// TIA Portal project "FK_PiPl" (V16)
// Lehrlingsprojekt

(* hardware
DEVICE "ET 200SP-Station_1"  ET 200SP-Station
   slot 0: "Baugruppenträger_0"  Rack  6ES5 710-8MAx1
   slot 1: "-20KF1"  CPU 1512SP F-1 PN  6ES7 512-1SK01-0AB0  V2.8
      slot 32768: "PROFINET-Schnittstelle_1"  X1
         slot 32771: "Port_3"  X1 P3
   slot 2: "-20KF5"  F-DI 8x24VDC HF  6ES7 136-6BA00-0CA0  V1.0
      slot 1: "-20KF5"  F-DI 8x24VDC HF
   slot 3: "-20KF6"  F-DQ 8x24VDC/0.5A PP HF  6ES7 136-6DC00-0CA0  V1.0
      slot 1: "-20KF6"  F-DQ 8x24VDC/0.5A PP HF
   slot 4: "-21KF1"  DI 16x24VDC ST  6ES7 131-6BH01-0BA0  V0.0
      slot 1: "-21KF1"  DI 16x24VDC ST
   slot 5: "-21KF4"  DQ 16x24VDC/0.5A ST  6ES7 132-6BH01-0BA0  V0.0
      slot 1: "-21KF4"  DQ 16x24VDC/0.5A ST
   slot 6: "-22KF1"  AI 2xU/I 2-,4-wire HS  6ES7 134-6HB00-0DA1  V2.0
      slot 1: "-22KF1"  AI 2xU/I 2-,4-wire HS
   slot 7: "-22KF3"  AQ 2xU ST  6ES7 135-6FB00-0BA1  V1.0
      slot 1: "-22KF3"  AQ 2xU ST
   slot 8: "Servermodul_1"  Server module  6ES7 193-6PA00-0AA0  V1.1
      slot 1: "Servermodul_1"  Server module
   slot 127: "BA 2xRJ45"  BA 2xRJ45  6ES7 193-6AR00-0AA0  V0.0
      slot 32769: "Port_1"  X1 P1  6ES7 193-6AR00-0AA0
      slot 32770: "Port_2"  X1 P2  6ES7 193-6AR00-0AA0
DEVICE "HMI_1"  KTP400 Comfort
   slot 0: "HMI_1"  KTP400 Comfort  6AV2 124-2DC01-0AX0  16.0.0.0
   slot 1: "HMI_RT_1"  KTP400 Comfort  6AV2 124-2DC01-0AX0  16.0.0.0
   slot 5: "HMI_1.IE_CP_1"  PROFINET Interface  16.0.0.0
      slot 1: "PROFINET Schnittstelle_1"  PROFINET Interface
         slot 1: "Port_1"  Port
   slot 7: "HMI_1.MPI/DP_CP_1"  MPI/DP Interface  16.0.0.0
*)

// ===== PLC "-20KF1"  CPU 1512SP F-1 PN =====
// protected blocks, not shown: "Datenbaustein_2", "Main_Safety_RTG1", "Main_Safety_RTG1_DB", "Safety_Variabeln"

VAR_GLOBAL   // PLC tag table "Standard-Variablentabelle"
   "Speicher_Start" AT %M4.0 : Bool;
   "Speicher_Vereinzelner" AT %M4.1 : Bool;
   "Speicher_Teil_Bereit" AT %M4.2 : Bool;
   "Flanke_Teil_Bereit" AT %M4.3 : Bool;
   "Deckel_Drauf" AT %M4.4 : Bool;
   "Sauger_an" AT %M4.6 : Bool;
   "Sauger_Runter" AT %M4.7 : Bool;
   "Schlitten_Ausfahren" AT %M5.0 : Bool;
   "Flanke_Schltten_Ausgefahren" AT %M5.1 : Bool;
   "Speicher_Schlitten_Ausgefahren" AT %M5.2 : Bool;
   "Flanke_Schlitten" AT %M5.3 : Bool;
   "Flanke_Teil" AT %M5.4 : Bool;
   "Speicher_Sauger_aktivierung" AT %M5.5 : Bool;
   "Teil_Fertig" AT %M5.6 : Bool;
   "Speicher_kein_Deckel" AT %M5.7 : Bool;
   "Start/Stop Auto" AT %M6.0 : Bool;
   "Flanke_Dekel" AT %M6.1 : Bool;
   "Merker_Flanke_kein_Deckel" AT %M6.2 : Bool;
   "Speicher_Rückstau" AT %M6.3 : Bool;
   "Förderband-vor_Speicher" AT %M4.5 : Bool;
   "Förderband_Zurück_Speicher" AT %M6.4 : Bool;
   "Start/Stop Hand" AT %M6.5 : Bool;
   "Druck_Sensor" AT %EW272 : Word;
   "Druck_Zwischenwert1" AT %MD100 : Real;
   "Druck_Zwischenwert2" AT %MD104 : Real;
   "Druck_Zwischenwert3" AT %MW108 : Int;
   "Druck_Zugross" AT %M6.6 : Bool;
   "Druck_Zuklein" AT %M6.7 : Bool;
   "Flanke p Man/Aut" AT %M7.0 : Bool;
   "Flanke n Man/Aut" AT %M7.1 : Bool;
   "Flanke Merker n Man/Aut" AT %M7.2 : Bool;
   "Flanke Merker p Man/Aut" AT %M7.3 : Bool;
   "Reset Man/Aut" AT %M7.4 : Bool;
END_VAR

VAR_GLOBAL   // PLC tag table "Systemflags"
   "System_Byte" AT %MB1 : Byte;   // Byte System
   "ME_PLC_First_Scan_Bit" AT %M1.0 : Bool;   // PLC First Scan Bit
   "ME_PLC_DiagStatusUpdate" AT %M1.1 : Bool;   // PLC Diagnostic Status Update
   "ME_PLC_TRUE" AT %M1.2 : Bool;   // PLC TRUE
   "ME_PLC_FALSE" AT %M1.3 : Bool;   // PLC FALSE
   "Clock_Byte" AT %MB50 : Byte;   // Byte PLC Clock
   "ME_PLC_Clock_0.1s" AT %M50.0 : Bool;   // PLC Clock 0.1s (10Hz )
   "ME_PLC_Clock_0.2s" AT %M50.1 : Bool;   // PLC Clock 0.2s (5Hz )
   "ME_PLC_Clock_0.4s" AT %M50.2 : Bool;   // PLC Clock 0.4s (2.5Hz )
   "ME_PLC_Clock_0.5s" AT %M50.3 : Bool;   // PLC Clock 0.5s (2Hz )
   "ME_PLC_Clock_0.8s" AT %M50.4 : Bool;   // PLC Clock 0.8s (1.25Hz )
   "ME_PLC_Clock_1.0s" AT %M50.5 : Bool;   // PLC Clock 1s (1Hz)
   "ME_PLC_Clock_1.6s" AT %M50.6 : Bool;   // PLC Clock 1.6s (0.625Hz )
   "ME_PLC_Clock_2.0s" AT %M50.7 : Bool;   // PLC Clock 2s (0.5Hz )
   "ME_PLC_FC_Test" AT %M2.0 : Bool;   // Testing Frequency Converters
   "ME_PLC_TRUE_to_do" AT %M2.2 : Bool;   // PLC TRUE to do
   "ME_PLC_FALSE_to_do" AT %M2.3 : Bool;   // PLC FALSE to do
   "ME_PLC_Led_Error" AT %M2.4 : Bool;   // PLC LED Error
   "ME_PLC_Led_Maint" AT %M2.5 : Bool;   // PLC LED Maintenance
   "ME_PLC_Startup_Rst" AT %M2.6 : Bool;   // PLC LED Startup Reset
   "ME_PLC_First_Scan_Bit_FC" AT %M2.1 : Bool;   // Call Frequency Converters
END_VAR

VAR_GLOBAL   // PLC tag table "IO-Pick&Placer"
   "CC_KF_FbEStop" AT %E0.0 : Bool;   // Rückmeldung Freigabe Not-Halt (81KF8)
   "PPTR_BG_InletPart" AT %E0.1 : Bool;   // Transportband Werkstück am Bandanfang (100BG1)
   "PPTR_BG_PartAtSep" AT %E0.2 : Bool;   // Transportband Werkstück am Vereinzeler (100BG2)
   "PPTR_BG_BackupPart" AT %E0.3 : Bool;   // Transportband Werkstück beim Bandende (100BG3)
   "PIPL_BG_CarrierRetracted" AT %E0.4 : Bool;   // Pick&Placer Schlitten eingefahren (120BG1)
   "PIPL_BG_CarrierExtended" AT %E0.5 : Bool;   // Pick&Placer Schlitten ausgefahren (120BG2)
   "PIPL_BG_SuctTop" AT %E0.6 : Bool;   // Pick&Placer Sauger oben (120BG3)
   "PIPL_BP_PartSuckedOn" AT %E0.7 : Bool;   // Pick&Placer Werkstück angesaugt (120PB4)
   "PIPL_Pa_SF_Reset" AT %E1.0 : Bool;   // Pick&Placer Bedienstelle Reset (160SF2)
   "PIPL_Pa_SF_Start" AT %E1.1 : Bool;   // Pick&Placer Bedienstelle Start (160SF3)
   "PIPL_Pa_SF_Stop" AT %E1.2 : Bool;   // Pick&Placer Bedienstelle Stop (160SF4)
   "PIPL_Pa_SF_ManAuto" AT %E1.3 : Bool;   // Pick&Placer Bedienstelle Manual - Auto (160SF5)
   "CC_Spare_I1.4" AT %E1.4 : Bool;   // Spare
   "CC_Spare_I1.5" AT %E1.5 : Bool;   // Spare
   "CC_Spare_I1.6" AT %E1.6 : Bool;   // Spare
   "CC_Spare_I1.7" AT %E1.7 : Bool;   // Spare
   "PPTR_MB_SeparatorExtend" AT %A0.0 : Bool;   // Transportband Vereinzeler ausfahren (105MB8)
   "PIPL_SC_Green" AT %A0.1 : Bool;   // Pick&Placer Turmleuchte grün (130PF1)
   "PIPL_SC_Yellow" AT %A0.2 : Bool;   // Pick&Placer Turmleuchte gelb (130PF1)
   "PIPL_SC_Red" AT %A0.3 : Bool;   // Pick&Placer Turmleuchte rot (130PF1)
   "PIPL_MB_CarrierExtend" AT %A0.4 : Bool;   // Pick&Placer Schlitten ausfahren (125MB1)
   "PIPL_MB_CarrierRetract" AT %A0.5 : Bool;   // Pick&Placer Schlitten einfahren (125MB2)
   "PIPL_MB_SuctDown" AT %A0.6 : Bool;   // Pick&Placer Sauger nach unten (125MB3)
   "PIPL_MB_VacuumOn" AT %A0.7 : Bool;   // Pick&Placer Vakuum ein (125MB4)
   "PIPL_Pa_PF_ControlCircuit" AT %A1.0 : Bool;   // Pick&Placer Bedienstelle LED Steuerspannung Ein (Reset) (160SF2)
   "PIPL_Pa_PF_Error" AT %A1.1 : Bool;   // Pick&Placer Bedienstelle LED Fehler (160PF2)
   "PIPL_Pa_PF_Start" AT %A1.2 : Bool;   // Pick&Placer Bedienstelle LED Start (160SF3)
   "CC_Spare_O1.3" AT %A1.3 : Bool;   // Spare
   "CC_Spare_O1.4" AT %A1.4 : Bool;   // Spare
   "CC_Spare_O1.5" AT %A1.5 : Bool;   // Spare
   "CC_Spare_O1.6" AT %A1.6 : Bool;   // Spare
   "CC_Spare_O1.7" AT %A1.7 : Bool;   // Spare
   "CC_Spare_IW274" AT %EW274 : Word;   // Spare
   "PPTR_TF_DriveSpeed" AT %AW272 : Word;   // Transportband Bandmotor Geschwindigkeit Option (105TF1)
   "CC_Spare_OW274" AT %AW274 : Word;   // Spare
END_VAR

VAR_GLOBAL   // PLC tag table "IO-Pick&Placer-Safety"
   "PIPL_Pa_EStopCh1" AT %E1000.0 : Bool;   // Pick&Placer Bedienstelle Not-Halt Channel 1 (160SF1)
   "CC_Spare_I1000.1" AT %E1000.1 : Bool;   // Spare
   "CC_Spare_I1000.2" AT %E1000.2 : Bool;   // Spare
   "CC_Spare_I1000.3" AT %E1000.3 : Bool;   // Spare
   "PIPL_Pa_EStopCh2" AT %E1000.4 : Bool;   // Pick&Placer Bedienstelle Not-Halt Channel 2 (160SF1)
   "CC_Spare_I1000.5" AT %E1000.5 : Bool;   // Spare
   "CC_Spare_I1000.6" AT %E1000.6 : Bool;   // Spare
   "CC_Spare_I1000.7" AT %E1000.7 : Bool;   // Spare
   "CC_KF_EStopCh1" AT %A1050.0 : Bool;   // Freigabe Not-Halt Channel 1 (81KF7)
   "CC_KF_EStopCh2" AT %A1050.1 : Bool;   // Freigabe Not-Halt Channel 2 (81KF8)
   "PPTR_TF_DriveForward" AT %A1050.2 : Bool;   // Transportband Bandmotor Vorwärts (105TF1)
   "PPTR_TF_DriveReverse" AT %A1050.3 : Bool;   // Transportband Bandmotor Rückwärts (105TF1)
   "CC_Spare_O1050.4" AT %A1050.4 : Bool;   // Spare
   "CC_Spare_O1050.5" AT %A1050.5 : Bool;   // Spare
   "CC_Spare_O1050.6" AT %A1050.6 : Bool;   // Spare
   "CC_Spare_O1050.7" AT %A1050.7 : Bool;   // Spare
END_VAR

DATA_BLOCK "HMI_Meldung"   // DB8
{ S7_Optimized_Access := 'FALSE' }
VERSION : 0.1
   VAR
      Druck_Wert_Gerundet : Int;
      Druck_Wert_genau : Real;
      Warnung : Struct
         "Not-Aus Quitieren" : Bool;   // Not-Aus Quitieren
         Rückstau : Bool;   // Rückstau
         Druck_Zugross : Bool;
         Druck_Zuklein : Bool;
         "4" : Bool;
         "5" : Bool;
         "6" : Bool;
         "7" : Bool;
         "10" : Bool;
         "11" : Bool;
         "12" : Bool;
         "13" : Bool;
         "14" : Bool;
         "15" : Bool;
         "16" : Bool;
         "17" : Bool;
      END_STRUCT;
      Fehler : Struct   // Triggerbit für Fehler
         "Deckel Fehlt" : Bool;   // Kein Deckel vorhanden
         "Not-Aus Betätigt" : Bool;   // Not-Aus lösen
         "2" : Bool;
         "3" : Bool;
         "4" : Bool;
         "5" : Bool;
         "6" : Bool;
         "7" : Bool;
         "10" : Bool;
         "11" : Bool;
         "12" : Bool;
         "13" : Bool;
         "14" : Bool;
         "15" : Bool;
         "16" : Bool;
         "17" : Bool;
      END_STRUCT;
      Meldungen : Struct
         "Werkstück erkannt" : Bool;   // Teil erkannt
         "1" : Bool;
         "2" : Bool;
         "3" : Bool;
         "4" : Bool;
         "5" : Bool;
         "6" : Bool;
         "7" : Bool;
         "10" : Bool;
         "11" : Bool;
         "12" : Bool;
         "13" : Bool;
         "14" : Bool;
         "15" : Bool;
         "16" : Bool;
         "17" : Bool;
      END_STRUCT;
   END_VAR
BEGIN
END_DATA_BLOCK

DATA_BLOCK "HMI_Variabeln"   // DB10
{ S7_Optimized_Access := 'TRUE' }
VERSION : 0.1
   VAR
      "Förderband vor" : Bool;
      "Förderbad Zurück" : Bool;
      "Schlitten Vor" : Bool;
      "Schlitten Zurück" : Bool;
      Sauger : Bool;
      LampenTest : Bool;
      "Sauger Runter" : Bool;
   END_VAR
BEGIN
END_DATA_BLOCK

DATA_BLOCK "Datenbaustein_1"   // DB122
{ S7_Optimized_Access := 'TRUE' }
VERSION : 0.1
   VAR
      Sammelstoerung : Bool;
      Lampe_Ein : Bool;
      Lampe_Aus : Bool;
      Reserve3 : Bool;
      Reserve4 : Bool;
      Reserve5 : Bool;
      Reserve6 : Bool;
      Reserve7 : Bool;
      Reserve8 : Bool;
      Reserve9 : Bool;
      Wert : Int;
      PIPL_Lamp_Red_Netflix : Bool;
   END_VAR
BEGIN
END_DATA_BLOCK

// folder: System blocks/Program resources

DATA_BLOCK "Verlängerung_Signal_Deckel"   // DB3
{ S7_Optimized_Access := 'TRUE' }
AUTHOR : Simatic
FAMILY : IEC
NAME : IEC_TMR
VERSION : 1.0
// stored: InstanceOfName IEC_TIMER
"IEC_TIMER"
BEGIN
END_DATA_BLOCK

DATA_BLOCK "Zeitverzögerung_Ausschalltung_Auto"   // DB5
{ S7_Optimized_Access := 'TRUE' }
AUTHOR : Simatic
FAMILY : IEC
NAME : IEC_TMR
VERSION : 1.0
// stored: InstanceOfName IEC_TIMER
"IEC_TIMER"
BEGIN
END_DATA_BLOCK

DATA_BLOCK "Rückstau"   // DB9
{ S7_Optimized_Access := 'TRUE' }
AUTHOR : Simatic
FAMILY : IEC
NAME : IEC_TMR
VERSION : 1.0
// stored: InstanceOfName IEC_TIMER
"IEC_TIMER"
BEGIN
END_DATA_BLOCK

DATA_BLOCK "Master_Reset"   // DB11
{ S7_Optimized_Access := 'TRUE' }
AUTHOR : Simatic
FAMILY : IEC
NAME : IEC_TMR
VERSION : 1.0
// stored: InstanceOfName IEC_TIMER
"IEC_TIMER"
BEGIN
END_DATA_BLOCK

DATA_BLOCK "Rückstau_Weg"   // DB12
{ S7_Optimized_Access := 'TRUE' }
AUTHOR : Simatic
FAMILY : IEC
NAME : IEC_TMR
VERSION : 1.0
// stored: InstanceOfName IEC_TIMER
"IEC_TIMER"
BEGIN
END_DATA_BLOCK

DATA_BLOCK "Kein_Deckel_Hand"   // DB13
{ S7_Optimized_Access := 'TRUE' }
AUTHOR : Simatic
FAMILY : IEC
NAME : IEC_TMR
VERSION : 1.0
// stored: InstanceOfName IEC_TIMER
"IEC_TIMER"
BEGIN
END_DATA_BLOCK

DATA_BLOCK "Kein_Deckel_Auto"   // DB14
{ S7_Optimized_Access := 'TRUE' }
AUTHOR : Simatic
FAMILY : IEC
NAME : IEC_TMR
VERSION : 1.0
// stored: InstanceOfName IEC_TIMER
"IEC_TIMER"
BEGIN
END_DATA_BLOCK

DATA_BLOCK "Zeitverzögerung_Ausschalltung_Hand"   // DB15
{ S7_Optimized_Access := 'TRUE' }
AUTHOR : Simatic
FAMILY : IEC
NAME : IEC_TMR
VERSION : 1.0
// stored: InstanceOfName IEC_TIMER
"IEC_TIMER"
BEGIN
END_DATA_BLOCK

// folder: (top level)

FUNCTION "Programm Auto" : Void   // FC1, FBD
{ S7_Optimized_Access := 'TRUE' }
VERSION : 0.1
   VAR_TEMP   // added for the SCL form of the ladder/FBD networks
      _w1 : Bool;
   END_VAR
BEGIN

REGION Network 1: SR des Starttasters
   // Wenn Starttaster gedrückt wird und ein Werkstück bereit steht zieht das SR
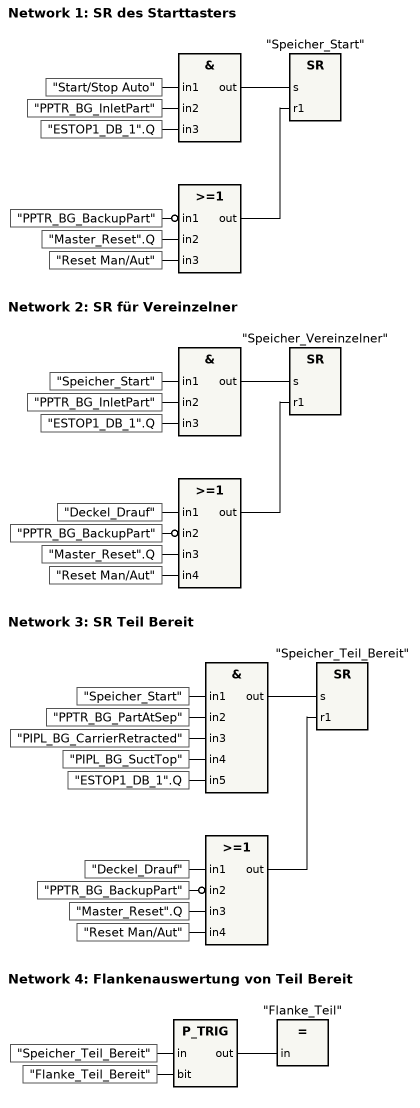
   IF "Start/Stop Auto" AND "PPTR_BG_InletPart" AND "ESTOP1_DB_1".Q THEN
       "Speicher_Start" := TRUE;   // SR flip-flop
   END_IF;
   IF NOT "PPTR_BG_BackupPart" OR "Master_Reset".Q OR "Reset Man/Aut" THEN "Speicher_Start" := FALSE; END_IF;
END_REGION

REGION Network 2: SR für Vereinzelner
   // Wenn das Programm gestartet wurde und das Werkstück auf dem Weg zum Vereinzelner ist zieht dieser an.
   IF "Speicher_Start" AND "PPTR_BG_InletPart" AND "ESTOP1_DB_1".Q THEN
       "Speicher_Vereinzelner" := TRUE;   // SR flip-flop
   END_IF;
   IF "Deckel_Drauf" OR NOT "PPTR_BG_BackupPart" OR "Master_Reset".Q OR "Reset Man/Aut" THEN
       "Speicher_Vereinzelner" := FALSE;
   END_IF;
END_REGION

REGION Network 3: SR Teil Bereit
   IF "Speicher_Start" AND "PPTR_BG_PartAtSep" AND "PIPL_BG_CarrierRetracted" AND "PIPL_BG_SuctTop" AND "ESTOP1_DB_1".Q THEN
       "Speicher_Teil_Bereit" := TRUE;   // SR flip-flop
   END_IF;
   IF "Deckel_Drauf" OR NOT "PPTR_BG_BackupPart" OR "Master_Reset".Q OR "Reset Man/Aut" THEN
       "Speicher_Teil_Bereit" := FALSE;
   END_IF;
END_REGION

REGION Network 4: Flankenauswertung von Teil Bereit
   #_w1 := "Speicher_Teil_Bereit" AND NOT "Flanke_Teil_Bereit";   // rising edge
   "Flanke_Teil_Bereit" := "Speicher_Teil_Bereit";
   "Flanke_Teil" := #_w1;
END_REGION

REGION Network 5: SR Sauger an
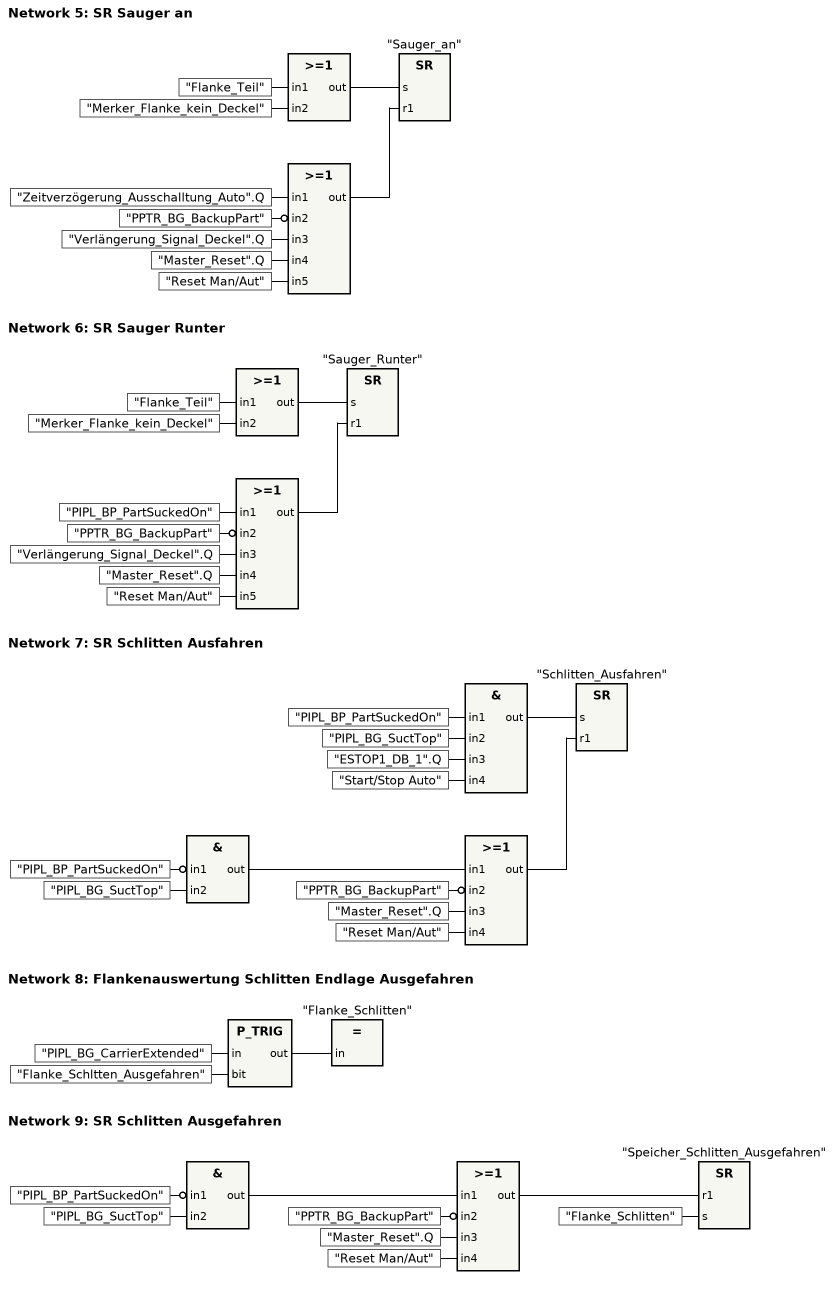
   IF "Flanke_Teil" OR "Merker_Flanke_kein_Deckel" THEN
       "Sauger_an" := TRUE;   // SR flip-flop
   END_IF;
   IF "Zeitverzögerung_Ausschalltung_Auto".Q OR NOT "PPTR_BG_BackupPart" OR "Verlängerung_Signal_Deckel".Q OR "Master_Reset".Q OR "Reset Man/Aut" THEN
       "Sauger_an" := FALSE;
   END_IF;
END_REGION

REGION Network 6: SR Sauger Runter
   IF "Flanke_Teil" OR "Merker_Flanke_kein_Deckel" THEN
       "Sauger_Runter" := TRUE;   // SR flip-flop
   END_IF;
   IF "PIPL_BP_PartSuckedOn" OR NOT "PPTR_BG_BackupPart" OR "Verlängerung_Signal_Deckel".Q OR "Master_Reset".Q OR "Reset Man/Aut" THEN
       "Sauger_Runter" := FALSE;
   END_IF;
END_REGION

REGION Network 7: SR Schlitten Ausfahren
   IF "PIPL_BP_PartSuckedOn" AND "PIPL_BG_SuctTop" AND "ESTOP1_DB_1".Q AND "Start/Stop Auto" THEN
       "Schlitten_Ausfahren" := TRUE;   // SR flip-flop
   END_IF;
   IF (NOT "PIPL_BP_PartSuckedOn" AND "PIPL_BG_SuctTop") OR NOT "PPTR_BG_BackupPart" OR "Master_Reset".Q OR "Reset Man/Aut" THEN
       "Schlitten_Ausfahren" := FALSE;
   END_IF;
END_REGION

REGION Network 8: Flankenauswertung Schlitten Endlage Ausgefahren
   #_w1 := "PIPL_BG_CarrierExtended" AND NOT "Flanke_Schltten_Ausgefahren";   // rising edge
   "Flanke_Schltten_Ausgefahren" := "PIPL_BG_CarrierExtended";
   "Flanke_Schlitten" := #_w1;
END_REGION

REGION Network 9: SR Schlitten Ausgefahren
   IF "Flanke_Schlitten" THEN
       "Speicher_Schlitten_Ausgefahren" := TRUE;   // SR flip-flop
   END_IF;
   IF (NOT "PIPL_BP_PartSuckedOn" AND "PIPL_BG_SuctTop") OR NOT "PPTR_BG_BackupPart" OR "Master_Reset".Q OR "Reset Man/Aut" THEN
       "Speicher_Schlitten_Ausgefahren" := FALSE;
   END_IF;
END_REGION

REGION Network 10: Zeitverzögerung für Saugerabschaltung
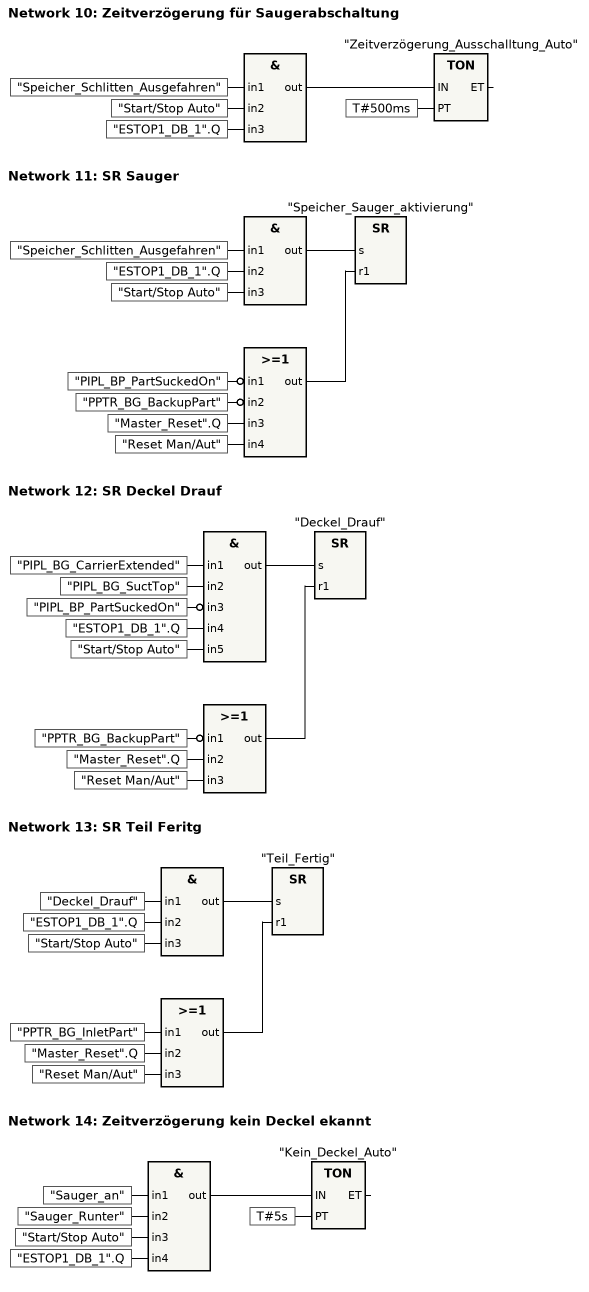
   "Zeitverzögerung_Ausschalltung_Auto".TON(IN := "Speicher_Schlitten_Ausgefahren" AND "Start/Stop Auto" AND "ESTOP1_DB_1".Q,
                           PT := T#500ms);
END_REGION

REGION Network 11: SR Sauger
   IF "Speicher_Schlitten_Ausgefahren" AND "ESTOP1_DB_1".Q AND "Start/Stop Auto" THEN
       "Speicher_Sauger_aktivierung" := TRUE;   // SR flip-flop
   END_IF;
   IF NOT "PIPL_BP_PartSuckedOn" OR NOT "PPTR_BG_BackupPart" OR "Master_Reset".Q OR "Reset Man/Aut" THEN
       "Speicher_Sauger_aktivierung" := FALSE;
   END_IF;
END_REGION

REGION Network 12: SR Deckel Drauf
   IF "PIPL_BG_CarrierExtended" AND "PIPL_BG_SuctTop" AND NOT "PIPL_BP_PartSuckedOn" AND "ESTOP1_DB_1".Q AND "Start/Stop Auto" THEN
       "Deckel_Drauf" := TRUE;   // SR flip-flop
   END_IF;
   IF NOT "PPTR_BG_BackupPart" OR "Master_Reset".Q OR "Reset Man/Aut" THEN "Deckel_Drauf" := FALSE; END_IF;
END_REGION

REGION Network 13: SR Teil Feritg
   IF "Deckel_Drauf" AND "ESTOP1_DB_1".Q AND "Start/Stop Auto" THEN
       "Teil_Fertig" := TRUE;   // SR flip-flop
   END_IF;
   IF "PPTR_BG_InletPart" OR "Master_Reset".Q OR "Reset Man/Aut" THEN "Teil_Fertig" := FALSE; END_IF;
END_REGION

REGION Network 14: Zeitverzögerung kein Deckel ekannt
   "Kein_Deckel_Auto".TON(IN := "Sauger_an" AND "Sauger_Runter" AND "Start/Stop Auto" AND "ESTOP1_DB_1".Q,
                          PT := T#5s);
END_REGION

REGION Network 15: SR kein Deckel
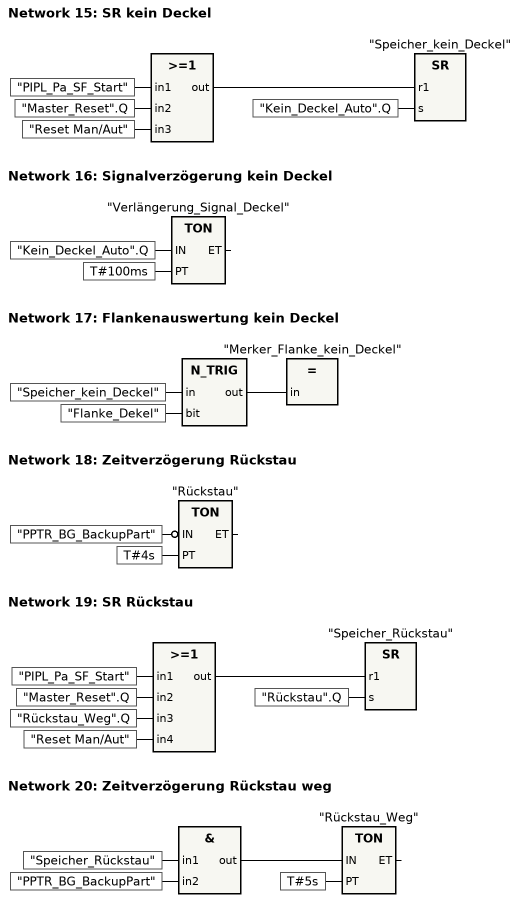
   IF "Kein_Deckel_Auto".Q THEN
       "Speicher_kein_Deckel" := TRUE;   // SR flip-flop
   END_IF;
   IF "PIPL_Pa_SF_Start" OR "Master_Reset".Q OR "Reset Man/Aut" THEN "Speicher_kein_Deckel" := FALSE; END_IF;
END_REGION

REGION Network 16: Signalverzögerung kein Deckel
   "Verlängerung_Signal_Deckel".TON(IN := "Kein_Deckel_Auto".Q, PT := T#100ms);
END_REGION

REGION Network 17: Flankenauswertung kein Deckel
   #_w1 := NOT "Speicher_kein_Deckel" AND "Flanke_Dekel";   // falling edge
   "Flanke_Dekel" := "Speicher_kein_Deckel";
   "Merker_Flanke_kein_Deckel" := #_w1;
END_REGION

REGION Network 18: Zeitverzögerung Rückstau
   "Rückstau".TON(IN := NOT "PPTR_BG_BackupPart", PT := T#4s);
END_REGION

REGION Network 19: SR Rückstau
   IF "Rückstau".Q THEN
       "Speicher_Rückstau" := TRUE;   // SR flip-flop
   END_IF;
   IF "PIPL_Pa_SF_Start" OR "Master_Reset".Q OR "Rückstau_Weg".Q OR "Reset Man/Aut" THEN
       "Speicher_Rückstau" := FALSE;
   END_IF;
END_REGION

REGION Network 20: Zeitverzögerung Rückstau weg
   "Rückstau_Weg".TON(IN := "Speicher_Rückstau" AND "PPTR_BG_BackupPart", PT := T#5s);
END_REGION
END_FUNCTION

FUNCTION "Start/Stop" : Void   // FC2, FBD
{ S7_Optimized_Access := 'TRUE' }
VERSION : 0.1
BEGIN

REGION Network 1: Start/Stop Hand
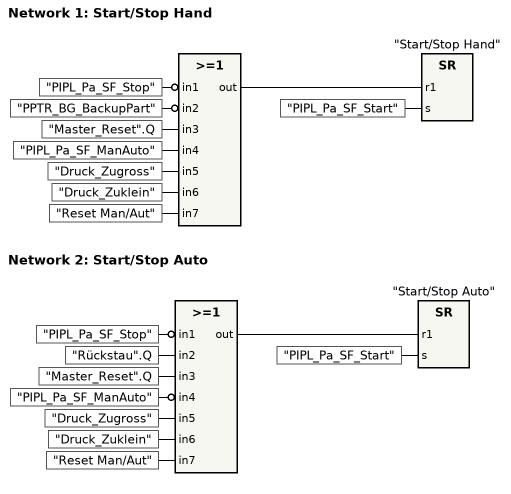
   IF "PIPL_Pa_SF_Start" THEN
       "Start/Stop Hand" := TRUE;   // SR flip-flop
   END_IF;
   IF NOT "PIPL_Pa_SF_Stop" OR NOT "PPTR_BG_BackupPart" OR "Master_Reset".Q OR "PIPL_Pa_SF_ManAuto" OR "Druck_Zugross" OR "Druck_Zuklein" OR "Reset Man/Aut" THEN
       "Start/Stop Hand" := FALSE;
   END_IF;
END_REGION

REGION Network 2: Start/Stop Auto
   IF "PIPL_Pa_SF_Start" THEN
       "Start/Stop Auto" := TRUE;   // SR flip-flop
   END_IF;
   IF NOT "PIPL_Pa_SF_Stop" OR "Rückstau".Q OR "Master_Reset".Q OR NOT "PIPL_Pa_SF_ManAuto" OR "Druck_Zugross" OR "Druck_Zuklein" OR "Reset Man/Aut" THEN
       "Start/Stop Auto" := FALSE;
   END_IF;
END_REGION
END_FUNCTION

FUNCTION "Master Reset" : Void   // FC3, FBD
{ S7_Optimized_Access := 'TRUE' }
VERSION : 0.1
   VAR_TEMP   // added for the SCL form of the ladder/FBD networks
      _w1 : Bool;
   END_VAR
BEGIN

REGION Network 1: Master Reset
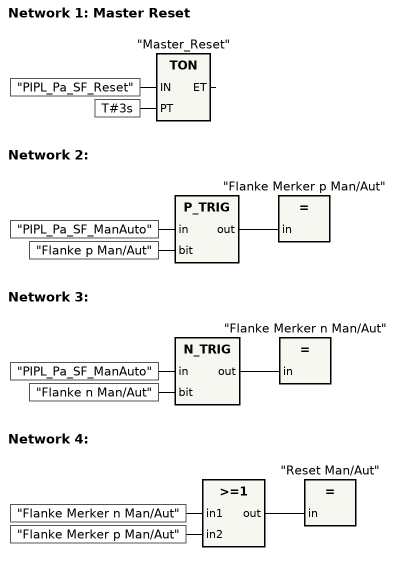
   "Master_Reset".TON(IN := "PIPL_Pa_SF_Reset", PT := T#3s);
END_REGION

REGION Network 2
   #_w1 := "PIPL_Pa_SF_ManAuto" AND NOT "Flanke p Man/Aut";   // rising edge
   "Flanke p Man/Aut" := "PIPL_Pa_SF_ManAuto";
   "Flanke Merker p Man/Aut" := #_w1;
END_REGION

REGION Network 3
   #_w1 := NOT "PIPL_Pa_SF_ManAuto" AND "Flanke n Man/Aut";   // falling edge
   "Flanke n Man/Aut" := "PIPL_Pa_SF_ManAuto";
   "Flanke Merker n Man/Aut" := #_w1;
END_REGION

REGION Network 4
   "Reset Man/Aut" := "Flanke Merker n Man/Aut" OR "Flanke Merker p Man/Aut";
END_REGION
END_FUNCTION

FUNCTION "Fehlermeldung" : Void   // FC4, FBD
{ S7_Optimized_Access := 'TRUE' }
VERSION : 0.1
BEGIN

REGION Network 1: Ausgang Fehlermeldung Rückstau
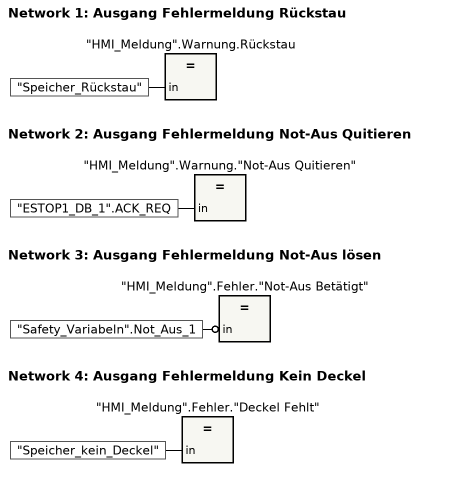
   "HMI_Meldung".Warnung.Rückstau := "Speicher_Rückstau";
END_REGION

REGION Network 2: Ausgang Fehlermeldung Not-Aus Quitieren
   "HMI_Meldung".Warnung."Not-Aus Quitieren" := "ESTOP1_DB_1".ACK_REQ;
END_REGION

REGION Network 3: Ausgang Fehlermeldung Not-Aus lösen
   "HMI_Meldung".Fehler."Not-Aus Betätigt" := NOT "Safety_Variabeln".Not_Aus_1;
END_REGION

REGION Network 4: Ausgang Fehlermeldung Kein Deckel
   "HMI_Meldung".Fehler."Deckel Fehlt" := "Speicher_kein_Deckel";
END_REGION
END_FUNCTION

FUNCTION "Programm Hand" : Void   // FC5, FBD
{ S7_Optimized_Access := 'TRUE' }
VERSION : 0.1
   VAR_TEMP   // added for the SCL form of the ladder/FBD networks
      _w1 : Bool;
   END_VAR
BEGIN

REGION Network 1: SR des Starttasters
   // Wenn Starttaster gedrückt wird und ein Werkstück bereit steht zieht das SR
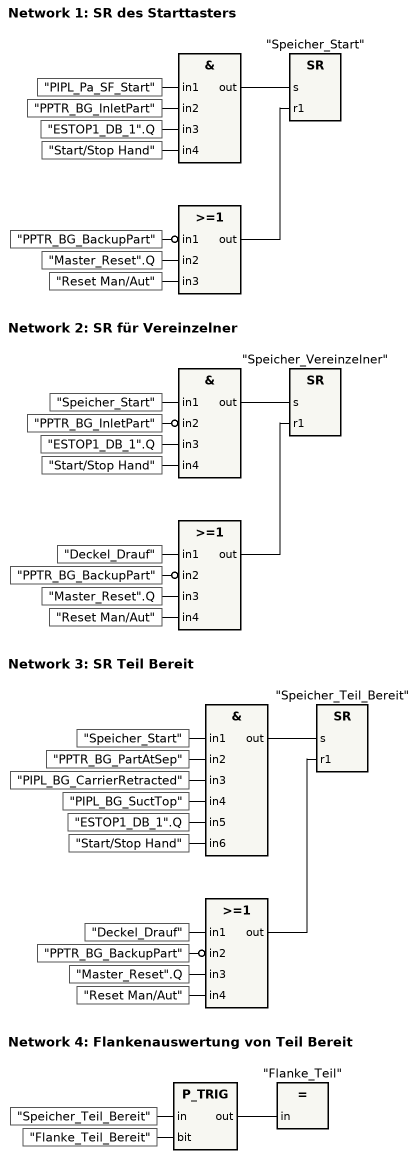
   IF "PIPL_Pa_SF_Start" AND "PPTR_BG_InletPart" AND "ESTOP1_DB_1".Q AND "Start/Stop Hand" THEN
       "Speicher_Start" := TRUE;   // SR flip-flop
   END_IF;
   IF NOT "PPTR_BG_BackupPart" OR "Master_Reset".Q OR "Reset Man/Aut" THEN "Speicher_Start" := FALSE; END_IF;
END_REGION

REGION Network 2: SR für Vereinzelner
   // Wenn das Programm gestartet wurde und das Werkstück auf dem Weg zum Vereinzelner ist zieht dieser an.
   IF "Speicher_Start" AND NOT "PPTR_BG_InletPart" AND "ESTOP1_DB_1".Q AND "Start/Stop Hand" THEN
       "Speicher_Vereinzelner" := TRUE;   // SR flip-flop
   END_IF;
   IF "Deckel_Drauf" OR NOT "PPTR_BG_BackupPart" OR "Master_Reset".Q OR "Reset Man/Aut" THEN
       "Speicher_Vereinzelner" := FALSE;
   END_IF;
END_REGION

REGION Network 3: SR Teil Bereit
   IF "Speicher_Start" AND "PPTR_BG_PartAtSep" AND "PIPL_BG_CarrierRetracted" AND "PIPL_BG_SuctTop" AND "ESTOP1_DB_1".Q AND "Start/Stop Hand" THEN
       "Speicher_Teil_Bereit" := TRUE;   // SR flip-flop
   END_IF;
   IF "Deckel_Drauf" OR NOT "PPTR_BG_BackupPart" OR "Master_Reset".Q OR "Reset Man/Aut" THEN
       "Speicher_Teil_Bereit" := FALSE;
   END_IF;
END_REGION

REGION Network 4: Flankenauswertung von Teil Bereit
   #_w1 := "Speicher_Teil_Bereit" AND NOT "Flanke_Teil_Bereit";   // rising edge
   "Flanke_Teil_Bereit" := "Speicher_Teil_Bereit";
   "Flanke_Teil" := #_w1;
END_REGION

REGION Network 5: SR Sauger Einschaltung